// TIA Portal project "Projeto caldeira - IHM" (V19)

(* hardware
DEVICE "SCALANCE X005"  SCALANCE X-Station
   slot 0: "SCALANCE X rack"  Rail
   slot 0: "Switch_1"  6GK5 005-0BA00-1AB2  V1.0
DEVICE "S7-1200 station_1"  S7-1200 Station
   slot 0: "Rack_0"  S7-1200 Rack  Rack  V1.0
   slot 1: "PLC_1"  CPU 1214C DC/DC/DC  6ES7 214-1AG40-0XB0  V4.6
DEVICE "HMI_1"  KTP600 Basic color PN
   slot 0: "HMI_1"  KTP600 Basic color PN  6AV6 647-0AD11-3AX0  12.0.0.0
   slot 1: "HMI_RT_1"  KTP600 Basic color PN  6AV6 647-0AD11-3AX0  12.0.0.0
   slot 5: "HMI_1.IE_CP_1"  PROFINET Interface  12.0.0.0
      slot 1: "PROFINET Interface_1"  PROFINET Interface
         slot 1: "Port_1"  Port
DEVICE "HMI_2"  KTP700 Basic PN
   slot 0: "HMI_2"  KTP700 Basic PN  6AV2 123-2GB03-0AX0  17.0.0.0
   slot 1: "HMI_RT_2"  KTP700 Basic PN  6AV2 123-2GB03-0AX0  17.0.0.0
   slot 5: "HMI_2.IE_CP_1"  PROFINET Interface  17.0.0.0
      slot 1: "PROFINET Interface_1"  PROFINET Interface
         slot 1: "Port_1"  Port
*)

// ===== PLC "PLC_1"  CPU 1214C DC/DC/DC =====

VAR_GLOBAL   // PLC tag table "Default tag table"
   "Motor" AT %I0.0 : Bool;
   "Turbina_!" AT %I0.1 : Bool;
   "Turbina_2" AT %I0.2 : Bool;
   "Tanque_1" AT %I0.3 : Bool;
   "Tanque_2" AT %I0.4 : Bool;
END_VAR

DATA_BLOCK "programação caldeira"   // DB1
{ S7_Optimized_Access := 'TRUE' }
VERSION : 0.1
   VAR
      Liga_caldeira : Bool;
      Liga_turbina : Bool;
      Liga_turbina_2 : Bool;
      Desliga_caldeira : Bool;
      Timer_1 : Bool;
      Timer_2 : Bool;
      Desliga : Bool;
      Liga : Bool;
   END_VAR
BEGIN
END_DATA_BLOCK

DATA_BLOCK "Lógica programação_DB"   // DB4
{ S7_Optimized_Access := 'TRUE' }
VERSION : 0.1
// stored: InstanceOfName Lógica programação
"Lógica programação"
BEGIN
END_DATA_BLOCK

DATA_BLOCK "Lógica programação_DB_1"   // DB5
{ S7_Optimized_Access := 'TRUE' }
VERSION : 0.1
// stored: InstanceOfName Lógica programação
"Lógica programação"
BEGIN
END_DATA_BLOCK

// folder: System blocks/Program resources

DATA_BLOCK "timer 1"   // DB2
{ S7_Optimized_Access := 'TRUE' }
AUTHOR : Simatic
FAMILY : IEC
NAME : IEC_TMR
VERSION : 1.0
// stored: InstanceOfName IEC_TIMER
"IEC_TIMER"
BEGIN
END_DATA_BLOCK

DATA_BLOCK "IEC_Timer_0_DB"   // DB3
{ S7_Optimized_Access := 'TRUE' }
AUTHOR : Simatic
FAMILY : IEC
NAME : IEC_TMR
VERSION : 1.0
// stored: InstanceOfName IEC_TIMER
"IEC_TIMER"
BEGIN
END_DATA_BLOCK

DATA_BLOCK "IEC_Timer_0_DB_1"   // DB6
{ S7_Optimized_Access := 'TRUE' }
AUTHOR : Simatic
FAMILY : IEC
NAME : IEC_TMR
VERSION : 1.0
// stored: InstanceOfName IEC_TIMER
"IEC_TIMER"
BEGIN
END_DATA_BLOCK

// folder: (top level)

FUNCTION_BLOCK "Lógica programação"   // FB1, LAD
{ S7_Optimized_Access := 'TRUE' }
VERSION : 0.1
BEGIN

REGION Network 1
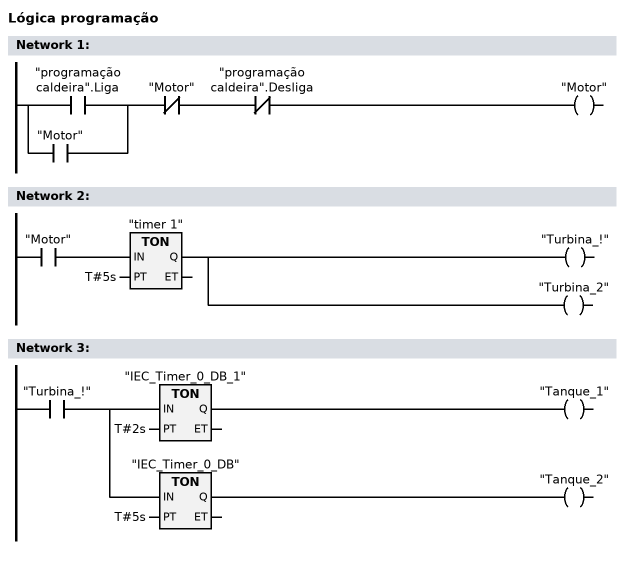
   RUNG wire#powerrail
      Contact( "programação caldeira".Liga )
      wire#w1
      I_Contact( "Motor" )
      I_Contact( "programação caldeira".Desliga )
      Coil( "Motor" )
   END_RUNG
   RUNG wire#powerrail
      Contact( "Motor" )
   END_RUNG wire#w1
   // the same network as SCL:
   "Motor" := ("programação caldeira".Liga OR "Motor") AND NOT "Motor" AND NOT "programação caldeira".Desliga;
END_REGION

REGION Network 2
   "timer 1".TON(IN := "Motor", PT := T#5s);
   "Turbina_!" := "timer 1".Q;
   "Turbina_2" := "timer 1".Q;
END_REGION

REGION Network 3
   "IEC_Timer_0_DB_1".TON(IN := "Turbina_!", PT := T#2s);
   "Tanque_1" := "IEC_Timer_0_DB_1".Q;
   "IEC_Timer_0_DB".TON(IN := "Turbina_!", PT := T#5s);
   "Tanque_2" := "IEC_Timer_0_DB".Q;
END_REGION
END_FUNCTION_BLOCK

ORGANIZATION_BLOCK "Main"   // OB1, LAD, ProgramCycle
TITLE = "Main Program Sweep (Cycle)"
{ S7_Optimized_Access := 'TRUE' }
VERSION : 0.1
   VAR_INPUT
      Initial_Call : Bool;   // Initial call of this OB
      Remanence : Bool;   // =True, if remanent data are available
   END_VAR
BEGIN

REGION Network 1
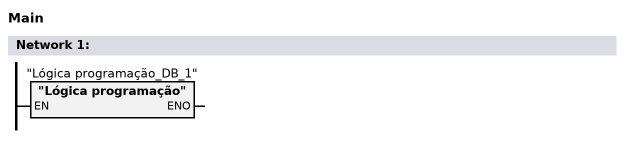
   RUNG wire#powerrail
      "Lógica programação_DB_1"()
   END_RUNG
   // the same network as SCL:
   "Lógica programação_DB_1"();   // "Lógica programação"
END_REGION
END_ORGANIZATION_BLOCK

(* ===== HMI "HMI_RT_1" =====
system functions are stored by id; their names below are inferred from use
connection "HMI_Connection_1": ETHERNET, SMART_S7_1200_OMS

HMI tags "Default tag table"
   "Tag_ScreenNumber" : UInt, internal
   "Turbina_!" : Bool = PLC Turbina_! AT %I0.1, 1 s
   "Turbina_2" : Bool = PLC Turbina_2 AT %I0.2, 1 s
   "Tanque_1" : Bool = PLC Tanque_1 AT %I0.3, 1 s
   "Tanque_2" : Bool = PLC Tanque_2 AT %I0.4, 1 s
   "programação caldeira_Liga_caldeira" : Bool = PLC "programação caldeira".Liga_caldeira, 1 s
   "Motor" : Bool = PLC Motor AT %I0.0, 1 s
   "programação caldeira_Desliga_caldeira" : Bool = PLC "programação caldeira".Desliga_caldeira, 1 s
   "programação caldeira_Liga" : Bool = PLC "programação caldeira".Liga, 1 s
   "programação caldeira_Desliga" : Bool = PLC "programação caldeira".Desliga, 1 s

Template "Template_1" 320x240
   Button "Exit" at 266,202 size 52x37; TextOff 'Exit'; PictureOff "ExitRuntime_KTP600_Basic_color_PN"; PictureOn "ExitRuntime_KTP600_Basic_color_PN"
      on Release: StopRuntime(0)
   Button "Template_Button" at 213,202 size 52x37; TextOff 'Text'
   Button "Template_Button_1" at 160,202 size 52x37; TextOff 'Text'
   Button "Template_Button_2" at 107,202 size 52x37; TextOff 'Text'
   Button "Template_Button_3" at 54,202 size 52x37; TextOff 'Text'
   Button "Start screen" at 1,202 size 52x37; TextOff 'Start screen'; PictureOff "NavigateHome_KTP600_Basic_color_PN"; PictureOn "NavigateHome_KTP600_Basic_color_PN"
      on Release: ActivateScreen("Root screen", 0)
   SymbolicIOField "Symbolic_IO_Field_Screen" at 69,7 size 164x24; TextOff '0'; TextOn '1'; TextList "TextList_ScreenNames"
      ProcessValue <- "Tag_ScreenNumber"
      on Change: ActivateScreenByNumber("Tag_ScreenNumber", 0)
   DateTimeField "HmiScreenItemData" at 235,19 size 85x19
   DateTimeField "HmiScreenItemData_1" at 235,0 size 85x19
   GraphicView "Logo" at 0,0 size 67x38; Picture "Logo of HMI_1"

screen "Root screen" 320x240, template "Template_1"
   on GenerateScreen: SetTag("Tag_ScreenNumber", 1)
   TextField "HmiScreenItemData" at 32,109 size 256x17; Text 'Welcome to HMI_1 (KTP600 Basic color PN)!'

screen "principal" 320x240
   TextField "Text field_1" at 76,6 size 186x29; Text 'Controle Caldeira'
   Button "Button_1" at 27,74 size 84x23; TextOff 'Liga'
      on Press: function_b14e0dd5("programação caldeira_Liga", 0)
   Circle "Circle_3" at 64,349 size 48x48
      Appearance <- "Turbina_2"
   Circle "Circle_4" at 0,349 size 48x48
      Appearance <- "Turbina_!"
   TextField "Text field_2" at 12,312 size 88x27; Text 'Turbinas'
   TextField "Text field_3" at 16,360 size 15x23; Text '1'
   TextField "Text field_4" at 80,361 size 15x23; Text '2'
   Rectangle "Rectangle_2" at 29,97 size 82x5
      Appearance <- "programação caldeira_Liga_caldeira"
   TextField "Text field_5" at 187,313 size 75x27; Text 'Válvula'
   Circle "Circle_1" at 345,347 size 48x48
      Appearance <- "Tanque_1"
   Circle "Circle_5" at 413,347 size 48x48
      Appearance <- "Tanque_2"
   TextField "Text field_6" at 364,315 size 75x27; Text 'Tanque'
   TextField "Text field_7" at 361,358 size 15x23; Text '1'
   TextField "Text field_8" at 429,359 size 15x23; Text '2'
   Circle "Circle_6" at 170,167 size 24x24
      Appearance <- "Turbina_2"
   Circle "Circle_7" at 139,166 size 24x24
      Appearance <- "Turbina_!"
   TextField "Text field_9" at 137,139 size 60x20; Text 'Turbinas'
   TextField "Text field_10" at 144,168 size 15x23; Text '1'
   TextField "Text field_11" at 175,168 size 15x22; Text '2'
   TextField "Text field_13" at 223,139 size 59x20; Text 'Tanques'
   Circle "Circle_9" at 222,168 size 24x24
      Appearance <- "Tanque_1"
   Circle "Circle_10" at 258,168 size 24x24
      Appearance <- "Tanque_2"
   TextField "Text field_14" at 227,169 size 15x23; Text '1'
   TextField "Text field_15" at 263,168 size 15x22; Text '2'
   Circle "Circle_8" at 39,165 size 21x21
      Appearance <- "Motor"
   TextField "Text field_12" at 28,139 size 44x20; Text 'Motor'
   Button "Button_2" at 198,74 size 84x23; TextOff 'Desliga'
      on Press: function_b14e0dd5("programação caldeira_Desliga", 0)
   Rectangle "Rectangle_3" at 200,97 size 82x5
      Appearance <- "programação caldeira_Desliga_caldeira"
*)

(* ===== HMI "HMI_RT_2" =====
system functions are stored by id; their names below are inferred from use
connection "HMI_Connection_2": ETHERNET, SMART_S7_1200_OMS

HMI tags "Default tag table"
   "Tag_ScreenNumber" : UInt, internal
   "programação caldeira_Liga" : Bool = PLC "programação caldeira".Liga, 1 s
   "programação caldeira_Desliga" : Bool = PLC "programação caldeira".Desliga, 1 s
   "Turbina_!" : Bool = PLC Turbina_! AT %I0.1, 1 s
   "Turbina_2" : Bool = PLC Turbina_2 AT %I0.2, 1 s
   "Motor" : Bool = PLC Motor AT %I0.0, 1 s
   "Tanque_1" : Bool = PLC Tanque_1 AT %I0.3, 1 s
   "Tanque_2" : Bool = PLC Tanque_2 AT %I0.4, 1 s

Template "Template_1" 800x480
   Button "Exit" at 714,429 size 71x50; TextOff 'Exit'; PictureOff "ExitRuntime_KTP700_Basic_PN_TR"; PictureOn "ExitRuntime_KTP700_Basic_PN_TR"
      on Release: StopRuntime(0)
   Button "Template_Button" at 614,429 size 71x50; TextOff 'Text'
   Button "Template_Button_1" at 514,429 size 71x50; TextOff 'Text'
   Button "Template_Button_2" at 414,429 size 71x50; TextOff 'Text'
   Button "Template_Button_3" at 314,429 size 71x50; TextOff 'Text'
   Button "Template_Button_4" at 214,429 size 71x50; TextOff 'Text'
   Button "Alarms" at 114,429 size 71x50; TextOff 'Alarms'; PictureOff "AlarmDisplay_KTP700_Basic_PN_TR"; PictureOn "AlarmDisplay_KTP700_Basic_PN_TR"
      on Release: function_ef3f5d25("Alarm window_Unacknowledged", -1)
   Button "Start screen" at 14,429 size 71x50; TextOff 'Start screen'; PictureOff "NavigateHome_KTP700_Basic_PN_TR"; PictureOn "NavigateHome_KTP700_Basic_PN_TR"
      on Release: ActivateScreen("Root screen", 0)
   SymbolicIOField "Symbolic_IO_Field_Screen" at 93,9 size 600x33; TextOff '0'; TextOn '1'; TextList "TextList_ScreenNames"
      ProcessValue <- "Tag_ScreenNumber"
      on Change: ActivateScreenByNumber("Tag_ScreenNumber", 0)
   DateTimeField "HmiScreenItemData" at 695,25 size 105x25
   DateTimeField "HmiScreenItemData_1" at 695,0 size 105x25
   GraphicView "Logo" at 0,0 size 91x51; Picture "Logo of HMI_2"

screen "Root screen" 800x480, template "Template_1"
   on GenerateScreen: SetTag("Tag_ScreenNumber", 1)
   TextField "HmiScreenItemData" at 80,225 size 640x25; Text 'Welcome to HMI_2 (KTP700 Basic+ PN)!'

screen "Screen_1" 800x480
   Button "Button_1" at 152,86 size 190x63; TextOff 'liga'
      on Click: SetBit("programação caldeira_Liga")
   Button "Button_2" at 485,91 size 187x56; TextOff 'desliga'
      on Click: SetBit("programação caldeira_Desliga")
   Rectangle "Rectangle_1" at 153,149 size 186x10
      Appearance <- "programação caldeira_Liga"
   Rectangle "Rectangle_2" at 485,148 size 186x10
      Appearance <- "programação caldeira_Desliga"
   TextField "Text field_1" at 165,220 size 78x27; Text 'Turbina'
   Circle "Circle_1" at 139,254 size 63x63
      Appearance <- "Turbina_!"
   Circle "Circle_2" at 213,257 size 63x63
      Appearance <- "Turbina_2"
   TextField "Text field_2" at 162,274 size 15x23; Text '1'
   TextField "Text field_3" at 238,275 size 15x23; Text '2'
   TextField "Text field_4" at 387,225 size 75x27; Text 'Tanque'
   Circle "Circle_3" at 358,252 size 63x63
      Appearance <- "Tanque_1"
   Circle "Circle_4" at 435,255 size 63x63
      Appearance <- "Tanque_2"
   TextField "Text field_5" at 382,272 size 15x23; Text '1'
   TextField "Text field_6" at 461,273 size 15x23; Text '2'
   TextField "Text field_7" at 577,227 size 62x27; Text 'Motor'
   Circle "Circle_5" at 575,258 size 63x63
      Appearance <- "Motor"
*)